// TIA Portal project "Urban Intersection Control System" (V17) (continued)
      R_Coil( "Traffic_Light_Operations_DB".MainStWest_Green )
      R_Coil( "Traffic_Light_Operations_DB".MainStWest_Yellow )
      R_Coil( "Traffic_Light_Operations_DB".MainStWest_Red )
   END_RUNG
   RUNG wire#powerrail
      R_Coil( "Traffic_Light_Operations_DB".CrossStSouth_Green )
      R_Coil( "Traffic_Light_Operations_DB".CrossStSouth_Yellow )
      R_Coil( "Traffic_Light_Operations_DB".CrossStSouth_Red )
      R_Coil( "Traffic_Light_Operations_DB".CrossStNorth_Green )
      R_Coil( "Traffic_Light_Operations_DB".CrossStNorth_Yellow )
      R_Coil( "Traffic_Light_Operations_DB".CrossStNorth_Red )
   END_RUNG
   // the same network as SCL:
   RESET_TIMER("MainStEast_Timer_DB");
   RESET_TIMER("MainStWest_Timer_DB");
   RESET_TIMER("CrossStSouth_Timer_DB");
   RESET_TIMER("CrossStNorth_Timer_DB");
   "Traffic_Light_Operations_DB".Initialize_Operation := FALSE;
   "Traffic_Light_Operations_DB".Traffic_Operations_Step := 0;
   "Traffic_Light_Operations_DB".MainStEast_Seconds := 0;
   "Traffic_Light_Operations_DB".MainStWest_Seconds := 0;
   "Traffic_Light_Operations_DB".CrossStSouth_Seconds := 0;
   "Traffic_Light_Operations_DB".CrossStNorth_Seconds := 0;
   "Traffic_Light_Operations_DB".MainStEast_Green := FALSE;
   "Traffic_Light_Operations_DB".MainStEast_Yellow := FALSE;
   "Traffic_Light_Operations_DB".MainStEast_Red := FALSE;
   "Traffic_Light_Operations_DB".MainStWest_Green := FALSE;
   "Traffic_Light_Operations_DB".MainStWest_Yellow := FALSE;
   "Traffic_Light_Operations_DB".MainStWest_Red := FALSE;
   "Traffic_Light_Operations_DB".CrossStSouth_Green := FALSE;
   "Traffic_Light_Operations_DB".CrossStSouth_Yellow := FALSE;
   "Traffic_Light_Operations_DB".CrossStSouth_Red := FALSE;
   "Traffic_Light_Operations_DB".CrossStNorth_Green := FALSE;
   "Traffic_Light_Operations_DB".CrossStNorth_Yellow := FALSE;
   "Traffic_Light_Operations_DB".CrossStNorth_Red := FALSE;
END_REGION

REGION Network 2: Pedestrian Status Reset
   // Resets the status of the pedestrian timers, pedestrian lights, and other variables
   RUNG wire#powerrail
      RT_Coil( "Ped_MainStEast_Timer_DB" )
      RT_Coil( "Ped_MainStWest_Timer_DB" )
      RT_Coil( "Ped_CrossStSouth_Timer_DB" )
      RT_Coil( "Ped_CrossStNorth_Timer_DB" )
   END_RUNG
   RUNG wire#powerrail
      R_Coil( "Pedestrian_Operations_DB".Walk_MainStEast )
      R_Coil( "Pedestrian_Operations_DB".Walk_MainStWest )
      R_Coil( "Pedestrian_Operations_DB".Walk_CrossStSouth )
      R_Coil( "Pedestrian_Operations_DB".Walk_CrossStNorth )
   END_RUNG
   RUNG wire#powerrail
      R_Coil( "Pedestrian_Operations_DB".DontWalk_MainStEast )
      R_Coil( "Pedestrian_Operations_DB".DontWalk_MainStWest )
      R_Coil( "Pedestrian_Operations_DB".DontWalk_CrossStSouth )
      R_Coil( "Pedestrian_Operations_DB".DontWalk_CrossStNorth )
   END_RUNG
   RUNG wire#powerrail
      Move(in := 0, out1 => "Pedestrian_Operations_DB".Ped_MainStEast_Seconds, out2 => "Pedestrian_Operations_DB".Ped_MainStWest_Seconds, out3 => "Pedestrian_Operations_DB".Ped_CrossStSouth_Seconds, out4 => "Pedestrian_Operations_DB".Ped_CrossStNorth_Seconds, out5 => "Pedestrian_Crossing_DB".PedCrossing_Seconds)
   END_RUNG
   RUNG wire#powerrail
      R_Coil( "Pedestrian_Operations_DB".Queue_MainStEast )
      R_Coil( "Pedestrian_Operations_DB".Queue_MainStWest )
      R_Coil( "Pedestrian_Operations_DB".Queue_CrossStSouth )
      R_Coil( "Pedestrian_Operations_DB".Queue_CrossStNorth )
   END_RUNG
   // the same network as SCL:
   RESET_TIMER("Ped_MainStEast_Timer_DB");
   RESET_TIMER("Ped_MainStWest_Timer_DB");
   RESET_TIMER("Ped_CrossStSouth_Timer_DB");
   RESET_TIMER("Ped_CrossStNorth_Timer_DB");
   "Pedestrian_Operations_DB".Walk_MainStEast := FALSE;
   "Pedestrian_Operations_DB".Walk_MainStWest := FALSE;
   "Pedestrian_Operations_DB".Walk_CrossStSouth := FALSE;
   "Pedestrian_Operations_DB".Walk_CrossStNorth := FALSE;
   "Pedestrian_Operations_DB".DontWalk_MainStEast := FALSE;
   "Pedestrian_Operations_DB".DontWalk_MainStWest := FALSE;
   "Pedestrian_Operations_DB".DontWalk_CrossStSouth := FALSE;
   "Pedestrian_Operations_DB".DontWalk_CrossStNorth := FALSE;
   "Pedestrian_Operations_DB".Ped_MainStEast_Seconds := 0;
   "Pedestrian_Operations_DB".Ped_MainStWest_Seconds := 0;
   "Pedestrian_Operations_DB".Ped_CrossStSouth_Seconds := 0;
   "Pedestrian_Operations_DB".Ped_CrossStNorth_Seconds := 0;
   "Pedestrian_Crossing_DB".PedCrossing_Seconds := 0;
   "Pedestrian_Operations_DB".Queue_MainStEast := FALSE;
   "Pedestrian_Operations_DB".Queue_MainStWest := FALSE;
   "Pedestrian_Operations_DB".Queue_CrossStSouth := FALSE;
   "Pedestrian_Operations_DB".Queue_CrossStNorth := FALSE;
END_REGION
END_FUNCTION_BLOCK

FUNCTION_BLOCK "Pedestrian_Operations"   // FB4, SCL
{ S7_Optimized_Access := 'TRUE' }
VERSION : 0.1
   VAR_INPUT
      PedPushButton_MainStEast : Bool;   // Push button for pedestrian crossing on eastern Main Street
      PedPushButton_MainStWest : Bool;   // Push button for pedestrian crossing on western Main Street
      PedPushButton_CrossStSouth : Bool;   // Push button for pedestrian crossing on southern Cross Street
      PedPushButton_CrossStNorth : Bool;   // Push button for pedestrian crossing on northern Cross Street
   END_VAR
   VAR_OUTPUT
      Walk_MainStEast : Bool;   // Pedestrian walk signal for eastern Main Street
      Walk_MainStWest : Bool;   // Pedestrian walk signal for western Main Street
      DontWalk_MainStEast : Bool;   // Pedestrian don't-walk signal for eastern Main Street
      DontWalk_MainStWest : Bool;   // Pedestrian don't-walk signal for western Main Street
      Walk_CrossStSouth : Bool;   // Pedestrian walk signal for southern Cross Street
      Walk_CrossStNorth : Bool;   // Pedestrian walk signal for northern Cross Street
      DontWalk_CrossStSouth : Bool;   // Pedestrian don't-walk signal for southern Cross Street
      DontWalk_CrossStNorth : Bool;   // Pedestrian don't-walk signal for northern Cross Street
      Queue_MainStEast : Bool;   // Pedestrian queue signal for eastern Main Street
      Queue_MainStWest : Bool;   // Pedestrian queue signal for western Main Street
      Queue_CrossStSouth : Bool;   // Pedestrian queue signal for southern Cross Street
      Queue_CrossStNorth : Bool;   // Pedestrian queue signal for northern Cross Street
   END_VAR
   VAR
      HMI_Ped_MainStEast_Command : Bool;   // Allows HMI to access push button for pedestrian crossing on eastern Main Street
      HMI_Ped_MainStWest_Command : Bool;   // Allows HMI to access push button for pedestrian crossing on western Main Street
      HMI_Ped_CrossStSouth_Command : Bool;   // Allows HMI to access push button for pedestrian crossing on southern Cross Street
      HMI_Ped_CrossStNorth_Command : Bool;   // Allows HMI to access push button for pedestrian crossing on northern Cross Street
      Ped_MainStEast_Seconds : Int;   // Allows HMI to read eastern Main Street pedestrian time
      Ped_MainStWest_Seconds : Int;   // Allows HMI to read western Main Street pedestrian time
      Ped_CrossStSouth_Seconds : Int;   // Allows HMI to read southern Cross Street pedestrian time
      Ped_CrossStNorth_Seconds : Int;   // Allows HMI to read northern Cross Street pedestrian time
      CrossingEnable_MainStEast : Bool;   // Pedestrian crossing has been granted for eastern Main Street
      CrossingEnable_MainStWest : Bool;   // Pedestrian crossing has been granted for western Main Street
      CrossingEnable_CrossStSouth : Bool;   // Pedestrian crossing has been granted for southern Cross Street
      CrossingEnable_CrossStNorth : Bool;   // Pedestrian crossing has been granted for northern Cross Street
   END_VAR
BEGIN
   (* ======= Pedestrian logic for eastern Main Street =======*)
   #CrossingEnable_MainStEast := "Traffic_Light_Operations_DB".MainStEast_Red AND "Traffic_Light_Operations_DB".MainStWest_Red;
   "Pedestrian_Crossing_DB"(PedPushButton := #PedPushButton_MainStEast,
                            Walk => #Walk_MainStEast,
                            DontWalk => #DontWalk_MainStEast,
                            Queue => #Queue_MainStEast,
                            PedCrossing_Seconds => #Ped_MainStEast_Seconds,
                            HMI_PedCrossing_Command := #HMI_Ped_MainStEast_Command,
                            CrossingEnable := #CrossingEnable_MainStEast);

   (* ======= Pedestrian logic for western Main Street =======*)
   #CrossingEnable_MainStWest := "Traffic_Light_Operations_DB".MainStWest_Red AND "Traffic_Light_Operations_DB".MainStEast_Red;
   "Pedestrian_Crossing_DB"(PedPushButton := #PedPushButton_MainStWest,
                            Walk => #Walk_MainStWest,
                            DontWalk => #DontWalk_MainStWest,
                            Queue => #Queue_MainStWest,
                            PedCrossing_Seconds => #Ped_MainStWest_Seconds,
                            HMI_PedCrossing_Command:= #HMI_Ped_MainStWest_Command,
                            CrossingEnable := #CrossingEnable_MainStWest);

   (* ======= Pedestrian logic for southern Cross Street =======*)
   #CrossingEnable_CrossStSouth := "Traffic_Light_Operations_DB".CrossStSouth_Red AND "Traffic_Light_Operations_DB".CrossStNorth_Red;
   "Pedestrian_Crossing_DB"(PedPushButton := #PedPushButton_CrossStSouth,
                            Walk => #Walk_CrossStSouth,
                            DontWalk => #DontWalk_CrossStSouth,
                            Queue => #Queue_CrossStSouth,
                            PedCrossing_Seconds => #Ped_CrossStSouth_Seconds,
                            HMI_PedCrossing_Command := #HMI_Ped_CrossStSouth_Command,
                            CrossingEnable := #CrossingEnable_CrossStSouth);

   (* ======= Pedestrian logic for northern Cross Street =======*)
   #CrossingEnable_CrossStNorth := "Traffic_Light_Operations_DB".CrossStNorth_Red AND"Traffic_Light_Operations_DB".CrossStSouth_Red;
   "Pedestrian_Crossing_DB"(PedPushButton := #PedPushButton_CrossStNorth,
                            Walk => #Walk_CrossStNorth,
                            DontWalk => #DontWalk_CrossStNorth,
                            Queue => #Queue_CrossStNorth,
                            PedCrossing_Seconds => #Ped_CrossStNorth_Seconds,
                            HMI_PedCrossing_Command := #HMI_Ped_CrossStNorth_Command,
                            CrossingEnable := #CrossingEnable_CrossStNorth);

   (*#Walk_MainStEast := FALSE;
   #DontWalk_MainStEast := TRUE;

   IF (#PedPushButton_MainStEast OR #HMI_Ped_MainStEast_Command) AND NOT #PedButton_Last THEN
       #Request := TRUE; (* Creates a request a pedestrian makes to cross *)
       #Queue_MainStEast := TRUE; (* Adds the request to the pedestrian queue until the red light appears *)
   END_IF;

   #PedButton_Last := #PedPushButton_MainStEast OR #HMI_Ped_MainStEast_Command;

   IF #Request AND "Traffic_Light_Operations_DB".MainStEast_Red = TRUE THEN
       (* Start timer *)
       "Ped_MainStEast_Timer_DB".TON(IN := TRUE, PT := T#8S); (*Pedestrian timer for eastern Main Street*) 
       #Ped_MainStEast_Seconds := DINT_TO_INT(TIME_TO_DINT("Ped_MainStEast_Timer_DB".ET) / 1000); (*Lets HMI read pedestrian time*)

       (* Walk phase active *)
       IF NOT "Ped_MainStEast_Timer_DB".Q THEN
           #Walk_MainStEast := TRUE;
           #DontWalk_MainStEast := FALSE;
           #Queue_MainStEast := FALSE; (*Resets the queue once it's safe to cross*)
       ELSE (* Time expired - return to Don't Walk *)
           #Walk_MainStEast := FALSE;
           #DontWalk_MainStEast := TRUE;
           #Request := FALSE; (* Crossing is done *)
       END_IF;
   ELSE (* Reset timer *)
       "Ped_MainStEast_Timer_DB".IN:= FALSE;
       #Ped_MainStEast_Seconds := 0;

       IF #Request AND NOT "Traffic_Light_Operations_DB".MainStEast_Red THEN
           #Queue_MainStEast := TRUE;  // still waiting
       END_IF;
   END_IF;
   (* ======================================================= *)

   (*Pedestrian logic for western Main Street*)
   #Walk_MainStWest := FALSE;
   #DontWalk_MainStWest := TRUE;
   IF (#PedPushButton_MainStWest OR #HMI_Ped_MainStWest_Command) AND "Traffic_Light_Operations_DB".MainStWest_Red = TRUE THEN
       "Ped_MainStWest_Timer_DB".TON(IN := TRUE, PT := T#8S); (*Pedestrian timer for western Main Street*)
       #Ped_MainStWest_Seconds := DINT_TO_INT(TIME_TO_DINT("Ped_MainStWest_Timer_DB".ET) / 1000);

       IF NOT "Ped_MainStWest_Timer_DB".Q THEN
           #Walk_MainStWest := TRUE;
           #DontWalk_MainStWest := FALSE;
       ELSE
           #Walk_MainStWest := FALSE;
           #DontWalk_MainStWest := TRUE;
       END_IF;

   ELSE
       "Ped_MainStWest_Timer_DB".IN := FALSE;
       #Ped_MainStWest_Seconds := 0;
   END_IF;



   (*Pedestrian logic for southern Cross Street*)
   #Walk_CrossStSouth := FALSE;
   #DontWalk_CrossStSouth := TRUE;
   IF (#PedPushButton_CrossStSouth OR #HMI_Ped_CrossStSouth_Command) AND "Traffic_Light_Operations_DB".CrossStSouth_Red = TRUE THEN
       "Ped_CrossStSouth_Timer_DB".TON(IN := TRUE, PT := T#8S); (*Pedestrian timer for southern Cross Street*)
       #Ped_CrossStSouth_Seconds := DINT_TO_INT(TIME_TO_DINT("Ped_CrossStSouth_Timer_DB".ET) / 1000);

       IF NOT "Ped_CrossStSouth_Timer_DB".Q THEN
           #Walk_CrossStSouth := TRUE;
           #DontWalk_CrossStSouth := FALSE;
       ELSE
           #Walk_CrossStSouth := FALSE;
           #DontWalk_CrossStSouth := TRUE;
       END_IF;

   ELSE
       "Ped_CrossStSouth_Timer_DB".IN := FALSE;
       #Ped_CrossStSouth_Seconds := 0;
   END_IF;

   (*Pedestrian logic for northern Cross Street*)
   #Walk_CrossStNorth := FALSE;
   #DontWalk_CrossStNorth := TRUE;
   IF (#PedPushButton_CrossStNorth OR #HMI_Ped_CrossStNorth_Command) AND "Traffic_Light_Operations_DB".CrossStNorth_Red = TRUE THEN
       "Ped_CrossStNorth_Timer_DB".TON(IN := TRUE, PT := T#8S); (*Pedestrian timer for northern Cross Street*)
       #Ped_CrossStNorth_Seconds := DINT_TO_INT(TIME_TO_DINT("Ped_CrossStNorth_Timer_DB".ET) / 1000);

       IF NOT "Ped_CrossStNorth_Timer_DB".Q THEN
           #Walk_CrossStNorth := TRUE;
           #DontWalk_CrossStNorth := FALSE;
       ELSE
           #Walk_CrossStNorth := FALSE;
           #DontWalk_CrossStNorth := TRUE;
       END_IF;

   ELSE
       "Ped_CrossStNorth_Timer_DB".IN := FALSE;
       #Ped_CrossStNorth_Seconds := 0;
   END_IF;*)
END_FUNCTION_BLOCK

FUNCTION_BLOCK "Pedestrian_Crossing"   // FB5, SCL
{ S7_Optimized_Access := 'TRUE' }
VERSION : 0.1
   VAR_INPUT
      CrossingEnable : Bool;   // Pedestrian crossing has been enabled
      PedPushButton : Bool;   // Set input for pedestrian push buttons
   END_VAR
   VAR_OUTPUT
      Walk : Bool;   // Set output for pedestrian walk signals
      DontWalk : Bool;   // Set output for pedestrian dont-walk signals
      Queue : Bool;   // Set output for queues
      PedCrossing_Seconds : Int;   // Set output for pedestrian time reading on HMI
   END_VAR
   VAR_IN_OUT
      HMI_PedCrossing_Command : Bool;   // Allows HMI to access push buttons for pedestrian crossing
   END_VAR
   VAR
      PedCrossing_Timer_Instance : TON_TIME;
      CrossingActive : Bool;   // Pedestrian crossing is active
      CrossingGranted : Bool;   // Pedestrian crossing has been granted
      PedButton_Last : Bool;   // Prevents multiple triggers when button is held
      Request : Bool;   // Creates a request a pedestrian makes to cross
   END_VAR
BEGIN
   #Walk := FALSE;
   #DontWalk := TRUE;

   IF (#PedPushButton OR #HMI_PedCrossing_Command) AND NOT #PedButton_Last THEN
       #Request := TRUE; (* Creates a request a pedestrian makes to cross *)
       #Queue := TRUE; (* Adds the request to the pedestrian queue until the red light appears *)
   END_IF;

   #PedButton_Last := #PedPushButton OR #HMI_PedCrossing_Command;

   IF #Request AND #CrossingEnable AND NOT #CrossingActive THEN
       #CrossingActive := TRUE;
       #Request := FALSE;
       #Queue := FALSE; (* Resets the queue once it's safe to cross *)
   END_IF;

   #PedCrossing_Timer_Instance.TON(IN := #CrossingActive, PT := T#8S); (* Pedestrian crossing timer *)
   #PedCrossing_Seconds := DINT_TO_INT(TIME_TO_DINT(#PedCrossing_Timer_Instance.ET) / 1000); (* Lets HMI read pedestrian time *)

   IF #CrossingActive THEN
       (*#PedCrossing_Timer_Instance.TON(IN := TRUE, PT := T#8S); (* Pedestrian crossing timer *)
       #PedCrossing_Seconds := DINT_TO_INT(TIME_TO_DINT(#PedCrossing_Timer_Instance.ET) / 1000); (* Lets HMI read pedestrian time *)*)
       (* Walk phase active *)
       #Walk := NOT #PedCrossing_Timer_Instance.Q;
       #DontWalk := #PedCrossing_Timer_Instance.Q;

       IF #PedCrossing_Timer_Instance.Q THEN (* Time expired - return to Don't Walk *)
           #CrossingActive := FALSE;
       END_IF;
   ELSE
        //#PedCrossing_Seconds := 0;
        #Walk := FALSE;
        #DontWalk := TRUE;

        IF #Request THEN 
            #Queue := TRUE;  // still waiting
        END_IF;
   END_IF;

       (*IF NOT #PedCrossing_Timer_Instance.Q THEN
           #Walk := TRUE;
           #DontWalk := FALSE;
           (*#Queue := FALSE; (* Resets the queue once it's safe to cross *)*)
       ELSE (* Time expired - return to Don't Walk *)
           #Walk := FALSE;
           #DontWalk := TRUE;
           #CrossingActive := FALSE;
           #Request := FALSE; (* Crossing is done *)
       END_IF;*)

   (*ELSE (* Reset timer *)
       (*#PedCrossing_Timer_Instance.IN := FALSE;*)
       #PedCrossing_Seconds := 0;

       IF #Request AND NOT #Red_Light THEN
           #Queue := TRUE;  // still waiting
       END_IF;*)
END_FUNCTION_BLOCK

ORGANIZATION_BLOCK "Main"   // OB1, LAD, ProgramCycle
TITLE = "Main Program Sweep (Cycle)"
{ S7_Optimized_Access := 'TRUE' }
VERSION : 0.1
   VAR_INPUT
      Initial_Call : Bool;   // Initial call of this OB
      Remanence : Bool;   // =True, if remanent data are available
   END_VAR
BEGIN

REGION Network 1: Main
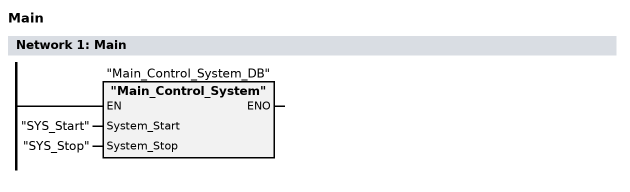
   RUNG wire#powerrail
      "Main_Control_System_DB"(System_Start := "SYS_Start", System_Stop := "SYS_Stop")
   END_RUNG
   // the same network as SCL:
   "Main_Control_System_DB"(System_Start := "SYS_Start", System_Stop := "SYS_Stop");   // "Main_Control_System"
END_REGION
END_ORGANIZATION_BLOCK

(* ===== HMI "HMI_RT_1" =====
system functions are stored by id; their names below are inferred from use
connection "HMI_Connection": ETHERNET, SMART_S7_1500_OMS

HMI tags "Default tag table"
   "Tag_ScreenNumber" : UInt, internal

HMI tags "UICS_HMI_Table"
   "MainStEast_RedLight" : Bool = PLC Traffic_Light_Operations_DB.MainStEast_Red AT %DB1.DBX0.0, 100 ms
   "MainStEast_YellowLight" : Bool = PLC Traffic_Light_Operations_DB.MainStEast_Yellow AT %DB1.DBX0.0, 100 ms
   "MainStEast_GreenLight" : Bool = PLC Traffic_Light_Operations_DB.MainStEast_Green AT %DB1.DBX0.0, 100 ms
   "MainStWest_RedLight" : Bool = PLC Traffic_Light_Operations_DB.MainStWest_Red AT %DB1.DBX0.0, 100 ms
   "MainStWest_YellowLight" : Bool = PLC Traffic_Light_Operations_DB.MainStWest_Yellow AT %DB1.DBX0.0, 100 ms
   "MainStWest_GreenLight" : Bool = PLC Traffic_Light_Operations_DB.MainStWest_Green AT %DB1.DBX0.0, 100 ms
   "CrossStSouth_RedLight" : Bool = PLC Traffic_Light_Operations_DB.CrossStSouth_Red AT %DB1.DBX0.0, 100 ms
   "CrossStSouth_YellowLight" : Bool = PLC Traffic_Light_Operations_DB.CrossStSouth_Yellow AT %DB1.DBX0.0, 100 ms
   "CrossStSouth_GreenLight" : Bool = PLC Traffic_Light_Operations_DB.CrossStSouth_Green AT %DB1.DBX0.0, 100 ms
   "CrossStNorth_RedLight" : Bool = PLC Traffic_Light_Operations_DB.CrossStNorth_Red AT %DB1.DBX0.0, 100 ms
   "CrossStNorth_YellowLight" : Bool = PLC Traffic_Light_Operations_DB.CrossStNorth_Yellow AT %DB1.DBX0.0, 100 ms
   "CrossStNorth_GreenLight" : Bool = PLC Traffic_Light_Operations_DB.CrossStNorth_Green AT %DB1.DBX0.0, 100 ms
   "MainStEast_Seconds" : Int = PLC Traffic_Light_Operations_DB.MainStEast_Seconds AT %DB1.DBX0.0, 100 ms
   "System_Running" : Bool = PLC Main_Control_System_DB.HMI_Run_Command AT %DB1.DBW0, 100 ms
   "Emergency_Stop" : Bool = PLC Main_Control_System_DB.Emergency_Stop AT %DB1.DBW0, 100 ms
   "Push_Button_Start" : Bool = PLC Main_Control_System_DB.HMI_Start_Command AT %DB1.DBX0.0, 100 ms
   "Push_Button_Stop" : Bool = PLC Main_Control_System_DB.HMI_Stop_Command AT %DB1.DBX0.0, 100 ms
   "CrossStNorth_Seconds" : Int = PLC Traffic_Light_Operations_DB.CrossStNorth_Seconds AT %DB1.DBW0, 100 ms
   "MainStWest_Seconds" : Int = PLC Traffic_Light_Operations_DB.MainStWest_Seconds AT %DB1.DBW0, 100 ms
   "CrossStSouth_Seconds" : Int = PLC Traffic_Light_Operations_DB.CrossStSouth_Seconds AT %DB1.DBW0, 100 ms
   "PedPushButton_MainStEast" : Bool = PLC Pedestrian_Operations_DB.HMI_Ped_MainStEast_Command AT %DB1.DBX0.0, 100 ms
   "PedPushButton_MainStWest" : Bool = PLC Pedestrian_Operations_DB.HMI_Ped_MainStWest_Command AT %DB1.DBX0.0, 100 ms
   "PedPushButton_CrossStSouth" : Bool = PLC Pedestrian_Operations_DB.HMI_Ped_CrossStSouth_Command AT %DB1.DBX0.0, 100 ms
   "PedPushButton_CrossStNorth" : Bool = PLC Pedestrian_Operations_DB.HMI_Ped_CrossStNorth_Command AT %DB1.DBX0.0, 100 ms
   "Walk_MainStEast" : Bool = PLC Pedestrian_Operations_DB.Walk_MainStEast AT %DB1.DBX0.0, 100 ms
   "Walk_MainStWest" : Bool = PLC Pedestrian_Operations_DB.Walk_MainStWest AT %DB1.DBX0.0, 100 ms
   "Walk_CrossStSouth" : Bool = PLC Pedestrian_Operations_DB.Walk_CrossStSouth AT %DB1.DBX0.0, 100 ms
   "Walk_CrossStNorth" : Bool = PLC Pedestrian_Operations_DB.Walk_CrossStNorth AT %DB1.DBX0.0, 100 ms
   "DontWalk_MainStEast" : Bool = PLC Pedestrian_Operations_DB.DontWalk_MainStEast AT %DB1.DBX0.0, 100 ms
   "DontWalk_MainStWest" : Bool = PLC Pedestrian_Operations_DB.DontWalk_MainStWest AT %DB1.DBX0.0, 100 ms
   "DontWalk_CrossStSouth" : Bool = PLC Pedestrian_Operations_DB.DontWalk_CrossStSouth AT %DB1.DBX0.0, 100 ms
   "DontWalk_CrossStNorth" : Bool = PLC Pedestrian_Operations_DB.DontWalk_CrossStNorth AT %DB1.DBX0.0, 100 ms
   "Ped_MainStEast_Seconds" : Int = PLC Pedestrian_Operations_DB.Ped_MainStEast_Seconds AT %DB1.DBX0.0, 100 ms
   "Ped_MainStWest_Seconds" : Int = PLC Pedestrian_Operations_DB.Ped_MainStWest_Seconds AT %DB1.DBX0.0, 100 ms
   "Ped_CrossStSouth_Seconds" : Int = PLC Pedestrian_Operations_DB.Ped_CrossStSouth_Seconds AT %DB1.DBX0.0, 100 ms
   "Ped_CrossStNorth_Seconds" : Int = PLC Pedestrian_Operations_DB.Ped_CrossStNorth_Seconds AT %DB1.DBX0.0, 100 ms
   "Ped_MainStEast_Queue" : Bool = PLC Pedestrian_Operations_DB.Queue_MainStEast AT %DB1.DBX0.0, 100 ms
   "Ped_MainStWest_Queue" : Bool = PLC Pedestrian_Operations_DB.Queue_MainStWest AT %DB1.DBX0.0, 100 ms
   "Ped_CrossStSouth_Queue" : Bool = PLC Pedestrian_Operations_DB.Queue_CrossStSouth AT %DB1.DBX0.0, 100 ms
   "Ped_CrossStNorth_Queue" : Bool = PLC Pedestrian_Operations_DB.Queue_CrossStNorth AT %DB1.DBX0.0, 100 ms

Template "Template_1" 1280x800
   Button "Exit" at 1182,752 size 67x47; TextOff 'Exit'; PictureOff "ExitRuntime_KTP1200_Basic_PN_TR"; PictureOn "ExitRuntime_KTP1200_Basic_PN_TR"
      on Release: StopRuntime(0)
   Button "Template_Button" at 1054,752 size 67x47; TextOff 'Text'
   Button "Template_Button_1" at 926,752 size 67x47; TextOff 'Text'
   Button "Template_Button_2" at 798,752 size 67x47; TextOff 'Text'
   Button "Template_Button_3" at 670,752 size 67x47; TextOff 'Text'
   Button "Template_Button_4" at 542,752 size 67x47; TextOff 'Text'
   Button "Template_Button_5" at 414,752 size 67x47; TextOff 'Text'
   Button "Template_Button_6" at 286,752 size 67x47; TextOff 'Text'
   Button "Alarms" at 158,752 size 67x47; TextOff 'Alarms'; PictureOff "AlarmDisplay_KTP1200_Basic_PN_TR"; PictureOn "AlarmDisplay_KTP1200_Basic_PN_TR"
      on Release: function_ef3f5d25("Alarm window_Unacknowledged", -1)
   Button "Start screen" at 30,752 size 67x47; TextOff 'Start screen'; PictureOff "NavigateHome_KTP1200_Basic_PN_TR"; PictureOn "NavigateHome_KTP1200_Basic_PN_TR"
      on Release: ActivateScreen("Root screen", 0)
   SymbolicIOField "Symbolic_IO_Field_Screen" at 87,9 size 1086x30; TextOff '0'; TextOn '1'; TextList "TextList_ScreenNames"
      ProcessValue <- "Tag_ScreenNumber"
      on Change: ActivateScreenByNumber("Tag_ScreenNumber", 0)
   DateTimeField "HmiScreenItemData" at 1175,24 size 105x24
   DateTimeField "HmiScreenItemData_1" at 1175,0 size 105x24
   GraphicView "Logo" at 0,0 size 85x48; Picture "Logo of HMI_1"

screen "Root screen" 1280x800, template "Template_1"
   on GenerateScreen: SetTag("Tag_ScreenNumber", 1)
   TextField "HmiScreenItemData" at 128,384 size 1024x27; Text 'Welcome to HMI_1 (KTP1200 Basic+ PN)!'

screen "Screen_1" 1280x800
   GraphicView "Four_Way_Road" at 319,94 size 612x612; Picture "Graphic_2"
   Group "MainStWest_TL" at 455,398 size 50x100
   Group "CrossStSouth_TL" at 622,509 size 100x50
   Group "CrossStNorth_TL" at 524,224 size 100x50
   IOField "I/O field_1" at 1049,403 size 96x32; FormatPattern s99; Unit  s
      ProcessValue <- "MainStEast_Seconds"
   Button "Start_Button" at 28,690 size 96x32; TextOff 'Start'
      on Press: InvertBit("Push_Button_Start")
   Button "Stop_Button" at 193,690 size 96x32; TextOff 'Stop'
      on Press: InvertBit("Push_Button_Stop")
   Switch "Pushbutton_Square_G" at 50,740 size 50x50; CaptionText 'Switch'; TextOff '0'; TextOn '1'; PictureOff "Pushbutton_Square_G_Off_256c"; PictureOn "Pushbutton_Square_G_On_256c"
      ProcessValue <- "System_Running"
   Switch "Pushbutton_Square_R" at 214,740 size 50x50; CaptionText 'Switch'; TextOff '0'; TextOn '1'; PictureOff "Pushbutton_Square_R_Off_256c"; PictureOn "Pushbutton_Square_R_On_256c"
      ProcessValue <- "Emergency_Stop"
   Group "MainStEast_TL" at 751,301 size 50x100
   IOField "I/O field_4" at 577,752 size 96x32; FormatPattern s99; Unit  s
      ProcessValue <- "CrossStSouth_Seconds"
   TextField "Text field_5" at 974,376 size 263x25; Text 'Eastern Main St Traffic Time'
   TextField "Text field_6" at 516,724 size 263x25; Text 'Southern Cross St Traffic Time'
   IOField "I/O field_2" at 97,400 size 96x32; FormatPattern s99; Unit  s
      ProcessValue <- "MainStWest_Seconds"
   TextField "Text field_1" at 32,372 size 263x25; Text 'Western Main St Traffic Time'
   IOField "I/O field_3" at 577,49 size 96x32; FormatPattern s99; Unit  s
      ProcessValue <- "CrossStNorth_Seconds"
   TextField "Text field_2" at 516,21 size 263x25; Text 'Northern Cross St Traffic Time'
   Button "PedPushButton_MainStEast" at 761,148 size 150x30; TextOff 'Request Walk'
      on Press: InvertBit("PedPushButton_MainStEast")
   TextField "Text field_3" at 766,110 size 145x25; Text 'Eastern Main St'
   TextField "Text field_4" at 750,193 size 47x25; Text 'Walk'
   TextField "Text field_7" at 828,194 size 99x25; Text 'Don't Walk'
   GraphicIOField "WalkSignal_MainStEast" at 755,225 size 50x50; PictureOn "PilotLight_Square_GN_On_256c"; PictureOff "PilotLight_Square_GN_Off_256c"
      ProcessValue <- "Walk_MainStEast"
   GraphicIOField "DontWalkSignal_MainStEast" at 854,224 size 50x50; PictureOff "PilotLight_Square_GN_Off_256c"; PictureOn "PilotLight_Square_GN_On_256c"
      ProcessValue <- "DontWalk_MainStEast"
   IOField "I/O field_5" at 1046,218 size 96x32; FormatPattern s99; Unit  s
      ProcessValue <- "Ped_MainStEast_Seconds"
   TextField "Text field_8" at 951,176 size 290x25; Text 'Eastern Main St Pedestrian Time'
   TextField "Text field_9" at 15,582 size 290x25; Text 'Western Main St Pedestrian Time'
   TextField "Text field_10" at 15,178 size 304x25; Text 'Northern Cross St Pedestrian Time'
   TextField "Text field_11" at 962,597 size 304x25; Text 'Southern Cross St Pedestrian Time'
   GraphicIOField "WalkSignal_CrossStNorth" at 340,225 size 50x50; PictureOff "PilotLight_Square_GN_Off_256c"; PictureOn "PilotLight_Square_GN_On_256c"
      ProcessValue <- "Walk_CrossStNorth"
   TextField "Text field_12" at 340,192 size 47x25; Text 'Walk'
   GraphicIOField "DontWalkSignal_CrossStNorth" at 431,224 size 50x50; PictureOn "PilotLight_Square_GN_On_256c"; PictureOff "PilotLight_Square_GN_Off_256c"
      ProcessValue <- "DontWalk_CrossStNorth"
   TextField "Text field_13" at 400,192 size 99x25; Text 'Don't Walk'
   TextField "Text field_14" at 338,110 size 174x25; Text 'Northern Cross St'
   Button "PedPushButton_CrossStNorth" at 340,149 size 150x30; TextOff 'Request Walk'
      on Press: InvertBit("PedPushButton_CrossStNorth")
   GraphicIOField "WalkSignal_MainStWest" at 340,530 size 50x50; PictureOn "PilotLight_Square_GN_On_256c"; PictureOff "PilotLight_Square_GN_Off_256c"
      ProcessValue <- "Walk_MainStWest"
   GraphicIOField "DontWalkSignal_MainStWest" at 430,528 size 50x50; PictureOff "PilotLight_Square_GN_Off_256c"; PictureOn "PilotLight_Square_GN_On_256c"
      ProcessValue <- "DontWalk_MainStWest"
   Button "PedPushButton_MainStWest" at 340,622 size 150x30; TextOff 'Request Walk'
      on Press: InvertBit("PedPushButton_MainStWest")
   TextField "Text field_15" at 344,666 size 158x25; Text 'Western Main St'
   TextField "Text field_16" at 336,592 size 47x25; Text 'Walk'
   TextField "Text field_17" at 403,590 size 99x25; Text 'Don't Walk'
   GraphicIOField "WalkSignal_CrossStSouth" at 756,526 size 50x50; PictureOn "PilotLight_Square_GN_On_256c"; PictureOff "PilotLight_Square_GN_Off_256c"
      ProcessValue <- "Walk_CrossStSouth"
   TextField "Text field_18" at 754,590 size 47x25; Text 'Walk'
   GraphicIOField "DontWalkSignal_CrossStSouth" at 850,526 size 50x50; PictureOff "PilotLight_Square_GN_Off_256c"; PictureOn "PilotLight_Square_GN_On_256c"
      ProcessValue <- "DontWalk_CrossStSouth"
   TextField "Text field_19" at 832,588 size 99x25; Text 'Don't Walk'
   Button "PedPushButton_CrossStSouth" at 763,622 size 150x30; TextOff 'Request Walk'
      on Press: InvertBit("PedPushButton_CrossStSouth")
   TextField "Text field_20" at 755,665 size 164x25; Text 'Southern Cross St'
   IOField "I/O field_6" at 104,616 size 96x32; FormatPattern s99; Unit  s
      ProcessValue <- "Ped_MainStWest_Seconds"
   IOField "I/O field_7" at 1068,630 size 96x32; FormatPattern s99; Unit  s
      ProcessValue <- "Ped_CrossStSouth_Seconds"
   IOField "I/O field_8" at 99,220 size 96x32; FormatPattern s99; Unit  s
      ProcessValue <- "Ped_CrossStNorth_Seconds"
   GraphicIOField "PedQueueSignal_MainStEast" at 964,112 size 50x50; PictureOff "PilotLight_Square_GN_Off_256c"; PictureOn "PilotLight_Square_GN_On_256c"
      ProcessValue <- "Ped_MainStEast_Queue"
   TextField "Text field_21" at 1023,112 size 198x25; Text 'Eastern Main St Queue'
   GraphicIOField "PedQueueSignal_MainStWest" at 23,528 size 50x50; PictureOn "PilotLight_Square_GN_On_256c"; PictureOff "PilotLight_Square_GN_Off_256c"
      ProcessValue <- "Ped_MainStWest_Queue"
   TextField "Text field_22" at 82,528 size 205x25; Text 'Western Main St Queue'
   GraphicIOField "PedQueueSignal_CrossStNorth" at 23,112 size 50x50; PictureOff "PilotLight_Square_GN_Off_256c"; PictureOn "PilotLight_Square_GN_On_256c"
      ProcessValue <- "Ped_CrossStNorth_Queue"
   TextField "Text field_23" at 83,112 size 217x25; Text 'Northern Cross St Queue'
   GraphicIOField "PedQueueSignal_CrossStSouth" at 951,528 size 50x50; PictureOff "PilotLight_Square_GN_Off_256c"; PictureOn "PilotLight_Square_GN_On_256c"
      ProcessValue <- "Ped_CrossStSouth_Queue"
   TextField "Text field_24" at 1010,528 size 219x25; Text 'Southern Cross St Queue'
   Circle "Green_East" at 763,370 size 26x26
      Appearance <- "MainStEast_GreenLight"
   Circle "Red_East" at 763,310 size 26x26
      Appearance <- "MainStEast_RedLight"
   Circle "Yellow_East" at 763,340 size 26x26
      Appearance <- "MainStEast_YellowLight"
   Circle "Red_West" at 467,407 size 26x26
      Appearance <- "MainStWest_RedLight"
   Circle "Yellow_West" at 467,437 size 26x26
      Appearance <- "MainStWest_YellowLight"
   Circle "Green_West" at 467,467 size 26x26
      Appearance <- "MainStWest_GreenLight"
   Circle "Red_South" at 687,521 size 26x26
      Appearance <- "CrossStSouth_RedLight"
   Circle "Yellow_South" at 657,521 size 26x26
      Appearance <- "CrossStSouth_YellowLight"
   Circle "Green_South" at 627,521 size 26x26
      Appearance <- "CrossStSouth_GreenLight"
   Circle "Red_North" at 589,236 size 26x26
      Appearance <- "CrossStNorth_RedLight"
   Circle "Yellow_North" at 559,236 size 26x26
      Appearance <- "CrossStNorth_YellowLight"
   Circle "Green_North" at 529,236 size 26x26
      Appearance <- "CrossStNorth_GreenLight"
*)